HMI tags "Default tag table"
   "phisical_DB_OUT_burning_t" : Int = PLC phisical_DB.OUT_burning_t, 1 s
   "phisical_DB_OUT_fluid_t" : Int = PLC phisical_DB.OUT_fluid_t, 1 s
   "phisical_DB_IN_gas_flow" : Int = PLC phisical_DB.IN_gas_flow, 1 s
   "phisical_DB_OUT_tank_presure" : Int = PLC phisical_DB.OUT_tank_presure, 1 s
   "phisical_DB_IN_pimp_speed" : Int = PLC phisical_DB.IN_pimp_speed, 1 s
   "phisical_DB_OUT_flow_speed" : Int = PLC phisical_DB.OUT_flow_speed, 1 s
   "phisical_DB_IN_pump_state" : Bool = PLC phisical_DB.IN_pump_state, 1 s
   "phisical_DB_IN_valve_state" : Bool = PLC phisical_DB.IN_valve_state, 1 s
   "phisical_DB_OUT_fire_state" : Bool = PLC phisical_DB.OUT_fire_state, 1 s
   "phisical_DB_OUT_pump_err" : Bool = PLC phisical_DB.OUT_pump_err, 1 s
   "phisical_DB_OUT_residential_heeting" : Bool = PLC phisical_DB.OUT_residential_heeting, 1 s
   "phisical_DB_pump_failure" : Bool = PLC phisical_DB.pump_failure, 1 s
   "phisical_DB_tank_failure" : Bool = PLC phisical_DB.tank_failure, 1 s
   "actuators_output_pimp_speed" : Int = PLC actuators_output.pimp_speed AT %DB9.DBW2, 1 s
   "actuators_output_gas_flow" : Int = PLC actuators_output.gas_flow AT %DB9.DBW0, 1 s
   "actuators_output_valve_state" : Bool = PLC actuators_output.valve_state AT %DB9.DBX4.0, 1 s
   "sensor_inputs_burning_temperature" : Int = PLC sensor_inputs.burning_temperature, 1 s
   "sensor_inputs_system_presure" : Int = PLC sensor_inputs.system_presure, 1 s
   "sensor_inputs_fluid_t" : Int = PLC sensor_inputs.fluid_t, 1 s
   "sensor_inputs_flow_speed" : Int = PLC sensor_inputs.flow_speed, 1 s
   "control_DB_temperature_setpoint" : Int = PLC control_DB.temperature_setpoint AT %DB6.DBW0, 1 s
   "control_DB_presure_err" : Bool = PLC control_DB.presure_err AT %DB6.DBX4.1, 1 s

screen "Screen_1" 1680x1050
   SymbolLibrary "Symbol library_1" at 26,257 size 55x156
   SymbolLibrary "Symbol library_2" at 53,290 size 68x123
   SymbolLibrary "Symbol library_3" at 96,355 size 57x58
   SymbolLibrary "Symbol library_8" at 362,417 size 152x276
   Group "Group" at 26,257 size 127x156
   Group "Group_2" at 85,246 size 80x87
   SymbolLibrary "Symbol library_11" at 251,605 size 364x41
   Group "Group_8" at 473,612 size 113x27
   Group "Group_9" at 277,612 size 63x27
   SymbolLibrary "Symbol library_5" at 605,427 size 105x351
   SymbolLibrary "Symbol library_29" at 602,335 size 112x120
      Visibility <- "phisical_DB_tank_failure"
   SymbolLibrary "Symbol library_30" at 605,457 size 106x147
      Visibility <- "phisical_DB_tank_failure"
   SymbolLibrary "Symbol library_12" at 287,902 size 304x120
   TextField "Text field_4" at 337,951 size 125x34; Text 'GAS Tank'
   SymbolLibrary "Symbol library_13" at 477,929 size 72x76
   SymbolLibrary "Symbol library_22" at 97,253 size 58x63
      Visibility <- "phisical_DB_OUT_residential_heeting"
   SymbolLibrary "Symbol library_24" at 85,246 size 80x87
      Visibility <- "phisical_DB_OUT_residential_heeting"
   SymbolLibrary "Symbol library_26" at 185,682 size 84x167
      Visibility <- "phisical_DB_pump_failure"
   SymbolLibrary "Symbol library_19" at 185,682 size 84x167
      Appearance <- "phisical_DB_OUT_pump_err"
      Visibility <- "phisical_DB_pump_failure"
   SymbolLibrary "Symbol library_28" at 175,612 size 87x71
      Visibility <- "phisical_DB_pump_failure"
   SymbolLibrary "Symbol library_7" at 175,612 size 87x71
      Appearance <- "phisical_DB_OUT_pump_err"
      Visibility <- "phisical_DB_pump_failure"
   SymbolLibrary "Symbol library_31" at 514,612 size 38x27
      Visibility <- "phisical_DB_tank_failure"
   SymbolLibrary "Symbol library_32" at 473,612 size 42x27
      Visibility <- "phisical_DB_tank_failure"
   SymbolLibrary "Symbol library_33" at 551,612 size 35x27
      Visibility <- "phisical_DB_tank_failure"
   SymbolLibrary "Symbol library_35" at 311,612 size 29x27
      Visibility <- "phisical_DB_tank_failure"
   SymbolLibrary "Symbol library_34" at 277,612 size 35x27
      Visibility <- "phisical_DB_tank_failure"
   SymbolLibrary "Symbol library_36" at 399,432 size 78x60
      Visibility <- "phisical_DB_tank_failure"
   SymbolLibrary "Symbol library_37" at 440,458 size 45x39
      Visibility <- "phisical_DB_tank_failure"
   SymbolLibrary "Symbol library_38" at 443,305 size 45x39
      Visibility <- "phisical_DB_tank_failure"
   SymbolLibrary "Symbol library_9" at 399,338 size 78x81
   Group "Group_1" at 362,417 size 152x276
   Group "Group_6" at 399,432 size 86x65
   Group "Group_3" at 185,682 size 84x167
   SymbolLibrary "Symbol library_25" at 151,770 size 145x41
      Visibility <- "phisical_DB_OUT_pump_err"
   SymbolLibrary "Symbol library_27" at 230,642 size 46x104
      Visibility <- "phisical_DB_pump_failure"
   Group "Group_5" at 175,612 size 87x71
   Group "Group_4" at 151,642 size 145x207
   Group "Group_7" at 362,305 size 152x388
   Group "Group_10" at 251,605 size 364x41
   SymbolLibrary "Symbol library_15" at 407,661 size 47x50
   Group "Group_13" at 151,612 size 145x237
   SymbolLibrary "Symbol library_6" at 114,612 size 63x54
      Appearance <- "phisical_DB_IN_valve_state"
   SymbolLibrary "Symbol library_4" at 67,584 size 49x83
   SymbolLibrary "Symbol library_23" at 644,501 size 120x42
   Group "Group_15" at 602,335 size 112x443
   TextField "Text field_3" at 56,904 size 131x22; Text 'Circulation pump'
   TextField "Text field_8" at 24,925 size 215x58; Text 'Creates flow in heating system. Can be damaged if run with closed valve longer than 10s.'
   Group "Group_24" at 18,897 size 225x90
   TextField "Text field_9" at 225,889 size 25x22; Text 'A1'
   TextField "Text field_7" at 590,803 size 132x22; Text 'Gas Flow Control'
   TextField "Text field_10" at 558,824 size 208x58; Text 'Controls amount of gas flowing in to burning chamber. Can be opened from 0 to 100%'
   Group "Group_26" at 552,796 size 225x90
   TextField "Text field_11" at 759,788 size 25x22; Text 'A2'
   TextField "Text field_13" at 322,444 size 25x22; Text 'A3'
   TextField "Text field_14" at 334,321 size 25x22; Text 'S1'
   TextField "Text field_17" at 753,244 size 25x22; Text 'S3'
   TextField "Text field_20" at 349,138 size 25x22; Text 'S2'
   TextField "Text field_23" at 754,112 size 25x22; Text 'S4'
   TextField "Text field_26" at 1615,624 size 25x22; Text 'A3'
   TextField "Text field_27" at 1601,126 size 25x22; Text 'A1'
   TextField "Text field_28" at 1608,365 size 25x22; Text 'A2'
   TextField "Text field_29" at 1100,823 size 25x22; Text 'S1'
   TextField "Text field_30" at 1100,576 size 25x22; Text 'S3'
   TextField "Text field_31" at 1098,388 size 25x22; Text 'S4'
   TextField "Text field_32" at 1096,159 size 25x22; Text 'S2'
   Rectangle "Rectangle_10" at 1176,792 size 475x69
      Visibility <- "control_DB_presure_err"
   SymbolLibrary "Symbol library_21" at 36,361 size 20x267
   Button "Button_1" at 1511,8 size 164x32; TextOff 'Open task manager'
      on Click: function_dfded056()
   SymbolLibrary "Symbol library_16" at 418,718 size 22x191
   SymbolLibrary "Symbol library_17" at 407,757 size 70x90
      Appearance <- "phisical_DB_OUT_fire_state"
   SymbolLibrary "Symbol library_18" at 403,110 size 146x253
      Visibility <- "phisical_DB_OUT_fire_state"
   SymbolLibrary "Symbol library_20" at 36,624 size 33x39
   Gauge "Gauge_2" at 865,68 size 193x193; UnitText 't'; CaptionText 'Burning temperature'
      ProcessValue <- "sensor_inputs_burning_temperature"
   Gauge "Gauge_3" at 877,728 size 188x188; UnitText 'l/min'; CaptionText 'Flow speed'
      ProcessValue <- "sensor_inputs_flow_speed"
   Gauge "Gauge_4" at 877,495 size 197x197; UnitText 't'; CaptionText 'Liquid t'
      ProcessValue <- "sensor_inputs_fluid_t"
   Slider "Slider_1" at 1459,339 size 116x230; Caption 'Set gas flow'
      ProcessValue <- "actuators_output_gas_flow"
   Gauge "Gauge_5" at 877,301 size 181x181; UnitText 'psi'; CaptionText 'Liquid presure'
      ProcessValue <- "sensor_inputs_system_presure"
   Slider "Slider_2" at 1453,83 size 114x230; Caption 'Set pump speed'
      ProcessValue <- "actuators_output_pimp_speed"
   Switch "Switch_2" at 1453,609 size 141x47; TextOn 'ON'; CaptionText 'Flow switch/valve'; TextOff 'OFF'
      ProcessValue <- "actuators_output_valve_state"
   Group "Group_11" at 251,305 size 364x406
   SymbolLibrary "Symbol library_10" at 378,559 size 116x98
      Visibility <- "phisical_DB_OUT_fire_state"
   Group "Group_12" at 26,246 size 139x167
   Group "Group_14" at 67,584 size 229x265
   SymbolLibrary "Symbol library_39" at 535,457 size 56x165
      Visibility <- "phisical_DB_tank_failure"
   Group "Group_16" at 287,902 size 304x120
   TextField "Text field_5" at 118,18 size 565x62; Text 'Heeting System SCADA'
   Group "Group_17" at 149,570 size 62x77
   Group "Group_18" at 91,664 size 107x224
   Group "Group_19" at 74,385 size 95x216
   Group "Group_21" at 443,795 size 108x50
   Group "Group_23" at 602,335 size 162x443
   SymbolLibrary "Symbol library_40" at 352,484 size 44x121
   Group "Group_20" at 363,262 size 29x240
   Group "Group_25" at 18,883 size 236x104
   Group "Group_22" at 719,317 size 39x202
   Group "Group_27" at 552,782 size 236x104
   TextField "Text field_6" at 168,462 size 154x22; Text 'Heating liquid valve'
   TextField "Text field_12" at 162,487 size 168x76; Text 'Heating liquid flow valve. When closed heat is not supplied to the residential buildings.'
   Group "Group_28" at 317,437 size 35x35
   TextField "Text field_1" at 186,333 size 143x22; Text 'Flow speed sensor'
   TextField "Text field_2" at 169,356 size 177x58; Text 'Monitors heating liquid flow speed in liters per minute (l/min)'
   Group "Group_29" at 329,314 size 35x35
   TextField "Text field_15" at 589,256 size 157x22; Text 'Temperature Sensor'
   TextField "Text field_16" at 569,279 size 199x22; Text 'Monitors temperature in tank.'
   Group "Group_30" at 748,237 size 35x35
   TextField "Text field_18" at 204,159 size 133x40; Text 'Burning Chamber Temperature'
   TextField "Text field_19" at 189,200 size 158x58; Text 'Monitors gas burning temperature. Depends on gas amount.'
   Group "Group_31" at 344,131 size 35x35
   TextField "Text field_21" at 609,124 size 120x22; Text 'Presure Sensor'
   TextField "Text field_22" at 573,147 size 169x76; Text 'Monitors presure in tank. If presure reaches 50 psi heating system can be damaged'
   Group "Group_32" at 749,105 size 35x35
   TextField "Text field_24" at 630,607 size 51x40; Text 'Liqiod Tank'
   TextField "Text field_25" at 29,224 size 128x22; Text 'Residential area'
   Group "Group_33" at 1610,617 size 35x35
   Group "Group_34" at 1595,119 size 35x35
   Group "Group_35" at 1602,358 size 35x35
   Group "Group_36" at 1095,816 size 35x35
   Group "Group_37" at 1095,569 size 35x35
   Group "Group_38" at 1093,381 size 35x35
   Group "Group_39" at 1091,152 size 35x35
   Slider "Slider_3" at 1226,237 size 207x230; Caption 'Set Desired liquid temperature'
      ProcessValue <- "control_DB_temperature_setpoint"
   TextField "Text field_33" at 1192,811 size 309x37; Text 'Presure Exceded Error'
      Visibility <- "control_DB_presure_err"
   Button "Button_2" at 1534,811 size 96x32; TextOff 'Reset'
      Visibility <- "control_DB_presure_err"
      on Click: InvertBit("control_DB_presure_err")
*)